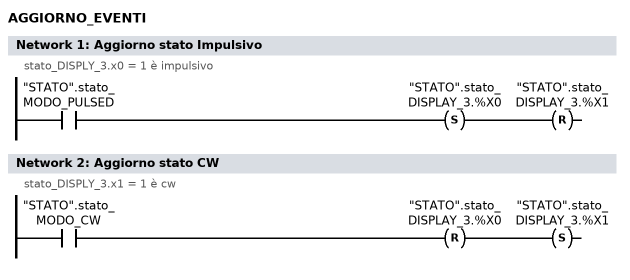
   RUNG wire#powerrail
      Contact( "STATO".stato_MODO_PULSED )
      S_Coil( "STATO".stato_DISPLAY_3.%X0 )
      R_Coil( "STATO".stato_DISPLAY_3.%X1 )
   END_RUNG
   // the same network as SCL:
   IF "STATO".stato_MODO_PULSED THEN
       "STATO".stato_DISPLAY_3.%X0 := TRUE;
       "STATO".stato_DISPLAY_3.%X1 := FALSE;
   END_IF;
END_REGION

REGION Network 2: Aggiorno stato CW
   // stato_DISPLY_3.x1 = 1 è cw
   RUNG wire#powerrail
      Contact( "STATO".stato_MODO_CW )
      R_Coil( "STATO".stato_DISPLAY_3.%X0 )
      S_Coil( "STATO".stato_DISPLAY_3.%X1 )
   END_RUNG
   // the same network as SCL:
   IF "STATO".stato_MODO_CW THEN
       "STATO".stato_DISPLAY_3.%X0 := FALSE;
       "STATO".stato_DISPLAY_3.%X1 := TRUE;
   END_IF;
END_REGION
END_FUNCTION

FUNCTION "LINEARIZZA_POTENZA" : Void   // FC11, LAD
TITLE = LINEARIZZA POTENZA
{ S7_Optimized_Access := 'FALSE' }
VERSION : 0.1
// Funzione di linearizzazione della potenza FWD e REFL
   VAR_TEMP   // added for the SCL form of the ladder/FBD networks
      _w1 : Bool;
   END_VAR
BEGIN

REGION Network 1: Calcolo indici N e N+1 tabella e punto adc&31
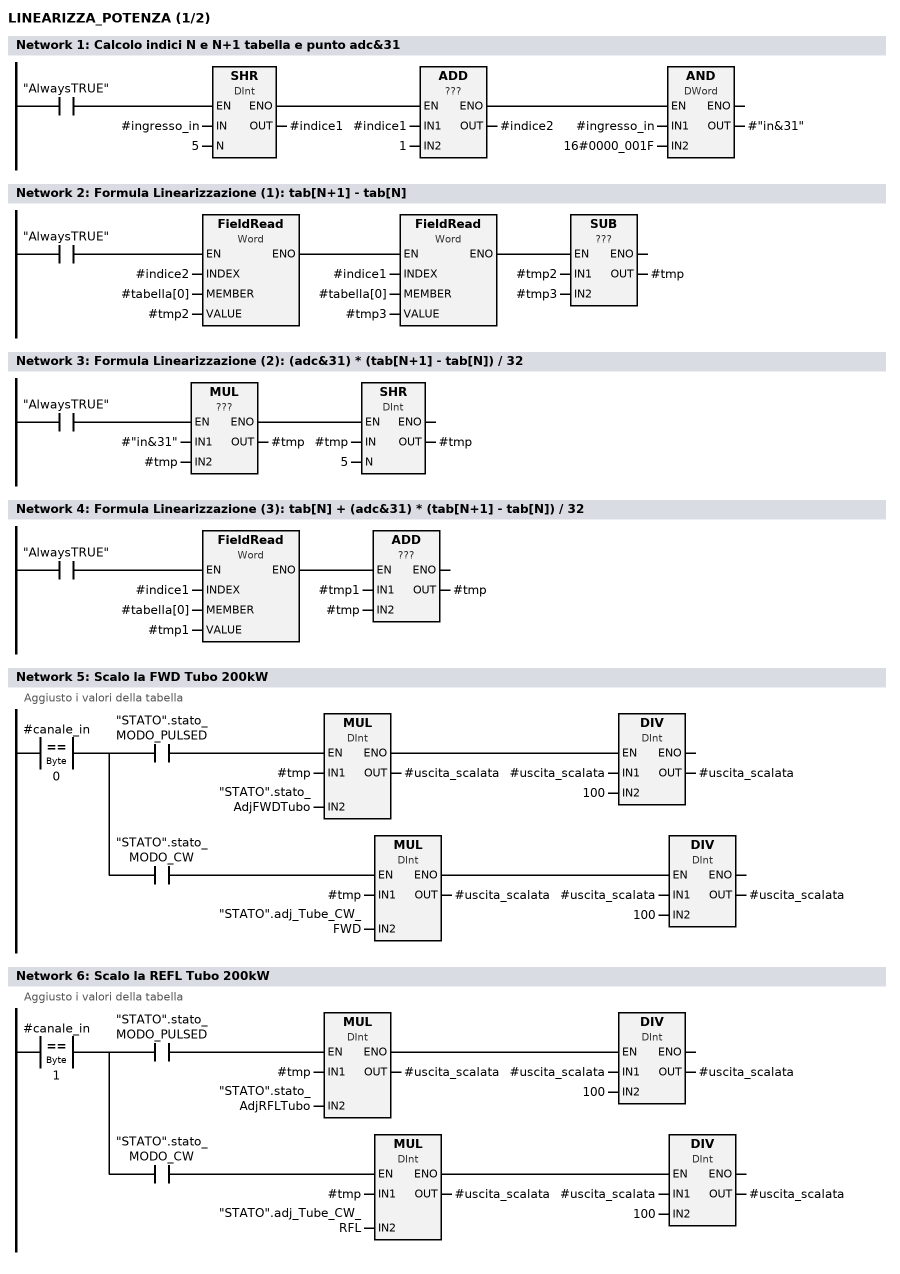
   // no checked SCL form for this network; see the picture
END_REGION

REGION Network 2: Formula Linearizzazione (1): tab[N+1] - tab[N]
   // no SCL statement known for FieldRead: written as a call
   // ENO of a box is taken as its EN; it also drops when the box reports an error
   #_w1 := "AlwaysTRUE";
   IF #_w1 THEN
       FieldRead(index := #indice2, member := #tabella[0], value := #tmp2);
       FieldRead(index := #indice1, member := #tabella[0], value := #tmp3);
       #tmp := #tmp2 - #tmp3;
   END_IF;
END_REGION

REGION Network 3: Formula Linearizzazione (2): (adc&31) * (tab[N+1] - tab[N]) / 32
   RUNG wire#powerrail
      Contact( "AlwaysTRUE" )
      { S7_Templates := "SrcType := ???" } Mul(in1 := #"in&31", in2 := #tmp, out => #tmp)
      { S7_Templates := "SrcType := DInt" } Shr(in := #tmp, n := 5, out => #tmp)
   END_RUNG
   // the same network as SCL:
   IF "AlwaysTRUE" THEN
       #tmp := #"in&31" * #tmp;
       #tmp := SHR(IN := #tmp, N := 5);
   END_IF;
END_REGION

REGION Network 4: Formula Linearizzazione (3): tab[N] + (adc&31) * (tab[N+1] - tab[N]) / 32
   // no SCL statement known for FieldRead: written as a call
   // ENO of a box is taken as its EN; it also drops when the box reports an error
   #_w1 := "AlwaysTRUE";
   IF #_w1 THEN
       FieldRead(index := #indice1, member := #tabella[0], value := #tmp1);
       #tmp := #tmp1 + #tmp;
   END_IF;
END_REGION

REGION Network 5: Scalo la FWD Tubo 200kW
   // Aggiusto i valori della tabella
   RUNG wire#powerrail
      { S7_Templates := "SrcType := Byte" } EQ_Contact(in1 := #canale_in, in2 := 0)
      wire#w1
      Contact( "STATO".stato_MODO_PULSED )
      { S7_Templates := "SrcType := DInt" } Mul(in1 := #tmp, in2 := "STATO".stato_AdjFWDTubo, out => #uscita_scalata)
      { S7_Templates := "SrcType := DInt" } Div(in1 := #uscita_scalata, in2 := 100, out => #uscita_scalata)
   END_RUNG
   RUNG wire#w1
      Contact( "STATO".stato_MODO_CW )
      { S7_Templates := "SrcType := DInt" } Mul(in1 := #tmp, in2 := "STATO".adj_Tube_CW_FWD, out => #uscita_scalata)
      { S7_Templates := "SrcType := DInt" } Div(in1 := #uscita_scalata, in2 := 100, out => #uscita_scalata)
   END_RUNG
   // the same network as SCL:
   #_w1 := #canale_in = 0;
   IF #_w1 AND "STATO".stato_MODO_PULSED THEN
       #uscita_scalata := #tmp * "STATO".stato_AdjFWDTubo;
       #uscita_scalata := #uscita_scalata / 100;
   END_IF;
   IF #_w1 AND "STATO".stato_MODO_CW THEN
       #uscita_scalata := #tmp * "STATO".adj_Tube_CW_FWD;
       #uscita_scalata := #uscita_scalata / 100;
   END_IF;
END_REGION

REGION Network 6: Scalo la REFL Tubo 200kW
   // Aggiusto i valori della tabella
   RUNG wire#powerrail
      { S7_Templates := "SrcType := Byte" } EQ_Contact(in1 := #canale_in, in2 := 1)
      wire#w1
      Contact( "STATO".stato_MODO_PULSED )
      { S7_Templates := "SrcType := DInt" } Mul(in1 := #tmp, in2 := "STATO".stato_AdjRFLTubo, out => #uscita_scalata)
      { S7_Templates := "SrcType := DInt" } Div(in1 := #uscita_scalata, in2 := 100, out => #uscita_scalata)
   END_RUNG
   RUNG wire#w1
      Contact( "STATO".stato_MODO_CW )
      { S7_Templates := "SrcType := DInt" } Mul(in1 := #tmp, in2 := "STATO".adj_Tube_CW_RFL, out => #uscita_scalata)
      { S7_Templates := "SrcType := DInt" } Div(in1 := #uscita_scalata, in2 := 100, out => #uscita_scalata)
   END_RUNG
   // the same network as SCL:
   #_w1 := #canale_in = 1;
   IF #_w1 AND "STATO".stato_MODO_PULSED THEN
       #uscita_scalata := #tmp * "STATO".stato_AdjRFLTubo;
       #uscita_scalata := #uscita_scalata / 100;
   END_IF;
   IF #_w1 AND "STATO".stato_MODO_CW THEN
       #uscita_scalata := #tmp * "STATO".adj_Tube_CW_RFL;
       #uscita_scalata := #uscita_scalata / 100;
   END_IF;
END_REGION

REGION Network 7: Scalo la FWD Stato Solido
   // Aggiusto i valori della tabella
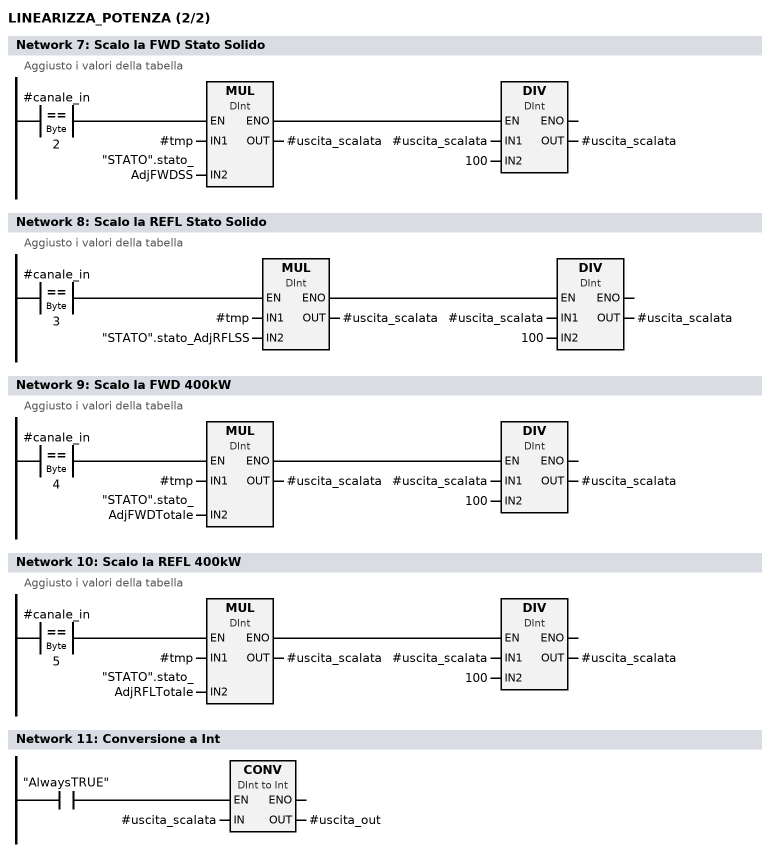
   RUNG wire#powerrail
      { S7_Templates := "SrcType := Byte" } EQ_Contact(in1 := #canale_in, in2 := 2)
      { S7_Templates := "SrcType := DInt" } Mul(in1 := #tmp, in2 := "STATO".stato_AdjFWDSS, out => #uscita_scalata)
      { S7_Templates := "SrcType := DInt" } Div(in1 := #uscita_scalata, in2 := 100, out => #uscita_scalata)
   END_RUNG
   // the same network as SCL:
   IF #canale_in = 2 THEN
       #uscita_scalata := #tmp * "STATO".stato_AdjFWDSS;
       #uscita_scalata := #uscita_scalata / 100;
   END_IF;
END_REGION

REGION Network 8: Scalo la REFL Stato Solido
   // Aggiusto i valori della tabella
   RUNG wire#powerrail
      { S7_Templates := "SrcType := Byte" } EQ_Contact(in1 := #canale_in, in2 := 3)
      { S7_Templates := "SrcType := DInt" } Mul(in1 := #tmp, in2 := "STATO".stato_AdjRFLSS, out => #uscita_scalata)
      { S7_Templates := "SrcType := DInt" } Div(in1 := #uscita_scalata, in2 := 100, out => #uscita_scalata)
   END_RUNG
   // the same network as SCL:
   IF #canale_in = 3 THEN
       #uscita_scalata := #tmp * "STATO".stato_AdjRFLSS;
       #uscita_scalata := #uscita_scalata / 100;
   END_IF;
END_REGION

REGION Network 9: Scalo la FWD 400kW
   // Aggiusto i valori della tabella
   RUNG wire#powerrail
      { S7_Templates := "SrcType := Byte" } EQ_Contact(in1 := #canale_in, in2 := 4)
      { S7_Templates := "SrcType := DInt" } Mul(in1 := #tmp, in2 := "STATO".stato_AdjFWDTotale, out => #uscita_scalata)
      { S7_Templates := "SrcType := DInt" } Div(in1 := #uscita_scalata, in2 := 100, out => #uscita_scalata)
   END_RUNG
   // the same network as SCL:
   IF #canale_in = 4 THEN
       #uscita_scalata := #tmp * "STATO".stato_AdjFWDTotale;
       #uscita_scalata := #uscita_scalata / 100;
   END_IF;
END_REGION

REGION Network 10: Scalo la REFL 400kW
   // Aggiusto i valori della tabella
   RUNG wire#powerrail
      { S7_Templates := "SrcType := Byte" } EQ_Contact(in1 := #canale_in, in2 := 5)
      { S7_Templates := "SrcType := DInt" } Mul(in1 := #tmp, in2 := "STATO".stato_AdjRFLTotale, out => #uscita_scalata)
      { S7_Templates := "SrcType := DInt" } Div(in1 := #uscita_scalata, in2 := 100, out => #uscita_scalata)
   END_RUNG
   // the same network as SCL:
   IF #canale_in = 5 THEN
       #uscita_scalata := #tmp * "STATO".stato_AdjRFLTotale;
       #uscita_scalata := #uscita_scalata / 100;
   END_IF;
END_REGION

REGION Network 11: Conversione a Int
   RUNG wire#powerrail
      Contact( "AlwaysTRUE" )
      { S7_Templates := "[SrcType := DInt, DestType := Int]" } Convert(in := #uscita_scalata, out => #uscita_out)
   END_RUNG
   // the same network as SCL:
   IF "AlwaysTRUE" THEN #uscita_out := DINT_TO_INT(#uscita_scalata); END_IF;
END_REGION
END_FUNCTION

FUNCTION "TRADUCI_TLS" : Void   // FC12, LAD
TITLE = TRADUCI_TLS
{ S7_Optimized_Access := 'FALSE' }
VERSION : 0.1
// Traduce gli stati/allarmi/misure in formato DATABLOCCO (EPICS_READ DB27) per l'invio al partner remoto EPICS.
   VAR_TEMP   // added for the SCL form of the ladder/FBD networks
      _w1 : Bool;
   END_VAR
BEGIN

REGION Network 1: Stato Locale/Remoto
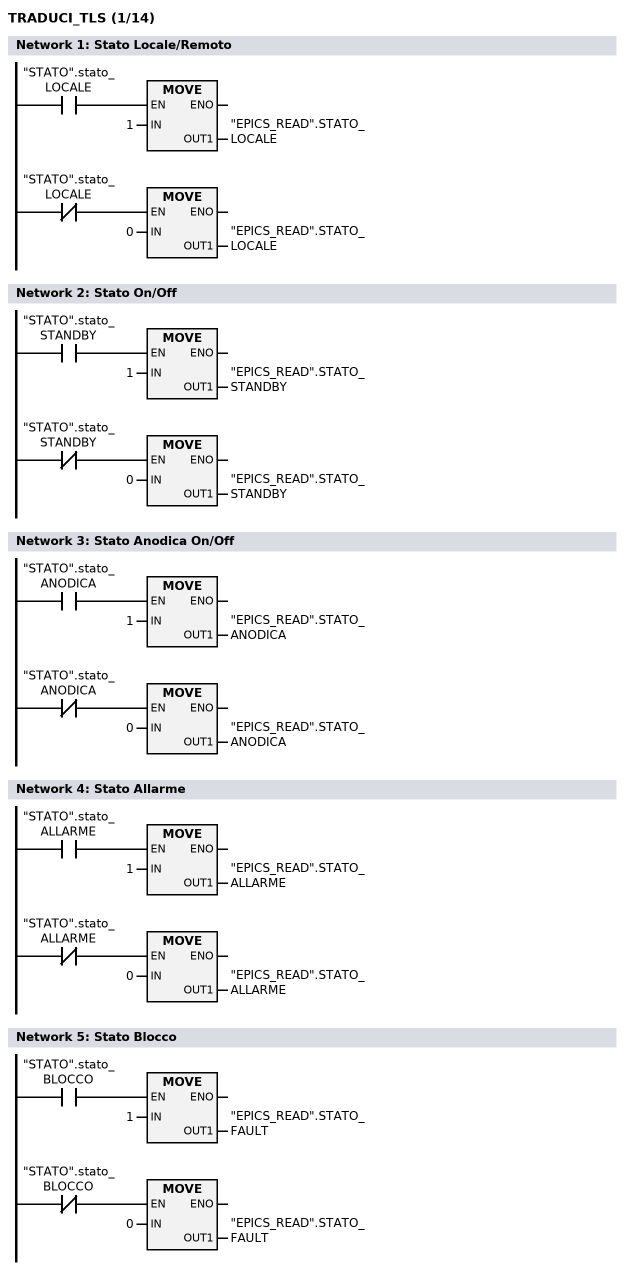
   RUNG wire#powerrail
      Contact( "STATO".stato_LOCALE )
      Move(in := 1, out1 => "EPICS_READ".STATO_LOCALE)
   END_RUNG
   RUNG wire#powerrail
      I_Contact( "STATO".stato_LOCALE )
      Move(in := 0, out1 => "EPICS_READ".STATO_LOCALE)
   END_RUNG
   // the same network as SCL:
   IF "STATO".stato_LOCALE THEN "EPICS_READ".STATO_LOCALE := 1; END_IF;
   IF NOT "STATO".stato_LOCALE THEN "EPICS_READ".STATO_LOCALE := 0; END_IF;
END_REGION

REGION Network 2: Stato On/Off
   RUNG wire#powerrail
      Contact( "STATO".stato_STANDBY )
      Move(in := 1, out1 => "EPICS_READ".STATO_STANDBY)
   END_RUNG
   RUNG wire#powerrail
      I_Contact( "STATO".stato_STANDBY )
      Move(in := 0, out1 => "EPICS_READ".STATO_STANDBY)
   END_RUNG
   // the same network as SCL:
   IF "STATO".stato_STANDBY THEN "EPICS_READ".STATO_STANDBY := 1; END_IF;
   IF NOT "STATO".stato_STANDBY THEN "EPICS_READ".STATO_STANDBY := 0; END_IF;
END_REGION

REGION Network 3: Stato Anodica On/Off
   RUNG wire#powerrail
      Contact( "STATO".stato_ANODICA )
      Move(in := 1, out1 => "EPICS_READ".STATO_ANODICA)
   END_RUNG
   RUNG wire#powerrail
      I_Contact( "STATO".stato_ANODICA )
      Move(in := 0, out1 => "EPICS_READ".STATO_ANODICA)
   END_RUNG
   // the same network as SCL:
   IF "STATO".stato_ANODICA THEN "EPICS_READ".STATO_ANODICA := 1; END_IF;
   IF NOT "STATO".stato_ANODICA THEN "EPICS_READ".STATO_ANODICA := 0; END_IF;
END_REGION

REGION Network 4: Stato Allarme
   RUNG wire#powerrail
      Contact( "STATO".stato_ALLARME )
      Move(in := 1, out1 => "EPICS_READ".STATO_ALLARME)
   END_RUNG
   RUNG wire#powerrail
      I_Contact( "STATO".stato_ALLARME )
      Move(in := 0, out1 => "EPICS_READ".STATO_ALLARME)
   END_RUNG
   // the same network as SCL:
   IF "STATO".stato_ALLARME THEN "EPICS_READ".STATO_ALLARME := 1; END_IF;
   IF NOT "STATO".stato_ALLARME THEN "EPICS_READ".STATO_ALLARME := 0; END_IF;
END_REGION

REGION Network 5: Stato Blocco
   RUNG wire#powerrail
      Contact( "STATO".stato_BLOCCO )
      Move(in := 1, out1 => "EPICS_READ".STATO_FAULT)
   END_RUNG
   RUNG wire#powerrail
      I_Contact( "STATO".stato_BLOCCO )
      Move(in := 0, out1 => "EPICS_READ".STATO_FAULT)
   END_RUNG
   // the same network as SCL:
   IF "STATO".stato_BLOCCO THEN "EPICS_READ".STATO_FAULT := 1; END_IF;
   IF NOT "STATO".stato_BLOCCO THEN "EPICS_READ".STATO_FAULT := 0; END_IF;
END_REGION

REGION Network 6: Impulsivo/CW
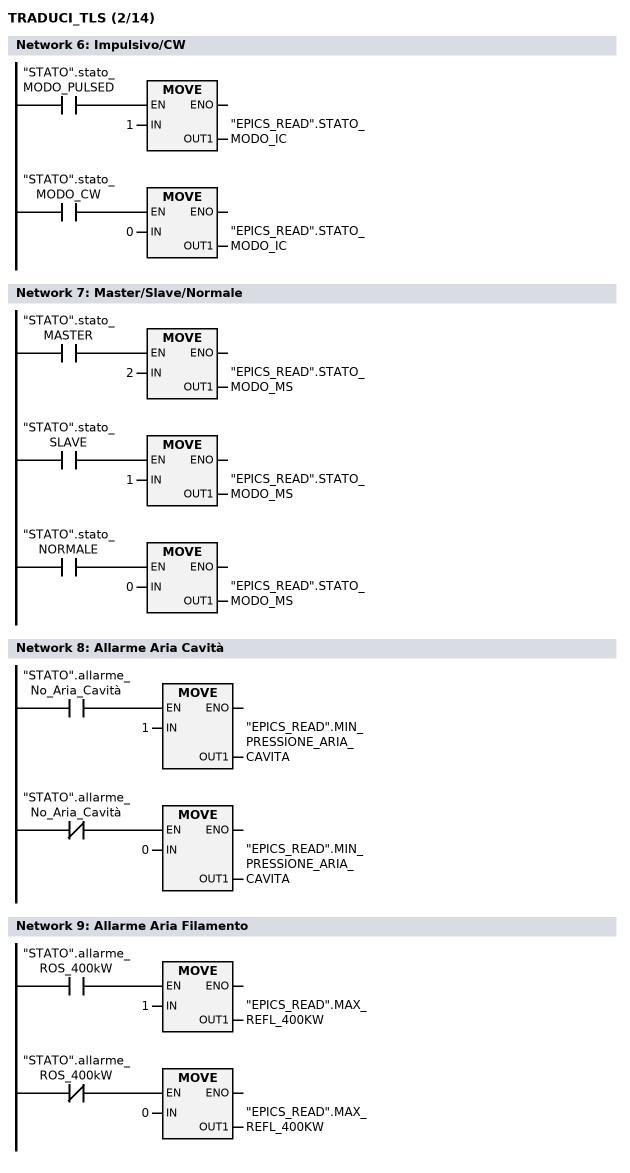
   RUNG wire#powerrail
      Contact( "STATO".stato_MODO_PULSED )
      Move(in := 1, out1 => "EPICS_READ".STATO_MODO_IC)
   END_RUNG
   RUNG wire#powerrail
      Contact( "STATO".stato_MODO_CW )
      Move(in := 0, out1 => "EPICS_READ".STATO_MODO_IC)
   END_RUNG
   // the same network as SCL:
   IF "STATO".stato_MODO_PULSED THEN "EPICS_READ".STATO_MODO_IC := 1; END_IF;
   IF "STATO".stato_MODO_CW THEN "EPICS_READ".STATO_MODO_IC := 0; END_IF;
END_REGION

REGION Network 7: Master/Slave/Normale
   RUNG wire#powerrail
      Contact( "STATO".stato_MASTER )
      Move(in := 2, out1 => "EPICS_READ".STATO_MODO_MS)
   END_RUNG
   RUNG wire#powerrail
      Contact( "STATO".stato_SLAVE )
      Move(in := 1, out1 => "EPICS_READ".STATO_MODO_MS)
   END_RUNG
   RUNG wire#powerrail
      Contact( "STATO".stato_NORMALE )
      Move(in := 0, out1 => "EPICS_READ".STATO_MODO_MS)
   END_RUNG
   // the same network as SCL:
   IF "STATO".stato_MASTER THEN "EPICS_READ".STATO_MODO_MS := 2; END_IF;
   IF "STATO".stato_SLAVE THEN "EPICS_READ".STATO_MODO_MS := 1; END_IF;
   IF "STATO".stato_NORMALE THEN "EPICS_READ".STATO_MODO_MS := 0; END_IF;
END_REGION

REGION Network 8: Allarme Aria Cavità
   RUNG wire#powerrail
      Contact( "STATO".allarme_No_Aria_Cavità )
      Move(in := 1, out1 => "EPICS_READ".MIN_PRESSIONE_ARIA_CAVITA)
   END_RUNG
   RUNG wire#powerrail
      I_Contact( "STATO".allarme_No_Aria_Cavità )
      Move(in := 0, out1 => "EPICS_READ".MIN_PRESSIONE_ARIA_CAVITA)
   END_RUNG
   // the same network as SCL:
   IF "STATO".allarme_No_Aria_Cavità THEN "EPICS_READ".MIN_PRESSIONE_ARIA_CAVITA := 1; END_IF;
   IF NOT "STATO".allarme_No_Aria_Cavità THEN "EPICS_READ".MIN_PRESSIONE_ARIA_CAVITA := 0; END_IF;
END_REGION

REGION Network 9: Allarme Aria Filamento
   RUNG wire#powerrail
      Contact( "STATO".allarme_ROS_400kW )
      Move(in := 1, out1 => "EPICS_READ".MAX_REFL_400KW)
   END_RUNG
   RUNG wire#powerrail
      I_Contact( "STATO".allarme_ROS_400kW )
      Move(in := 0, out1 => "EPICS_READ".MAX_REFL_400KW)
   END_RUNG
   // the same network as SCL:
   IF "STATO".allarme_ROS_400kW THEN "EPICS_READ".MAX_REFL_400KW := 1; END_IF;
   IF NOT "STATO".allarme_ROS_400kW THEN "EPICS_READ".MAX_REFL_400KW := 0; END_IF;
END_REGION

REGION Network 10: Allarme Flusso LQD Tubo
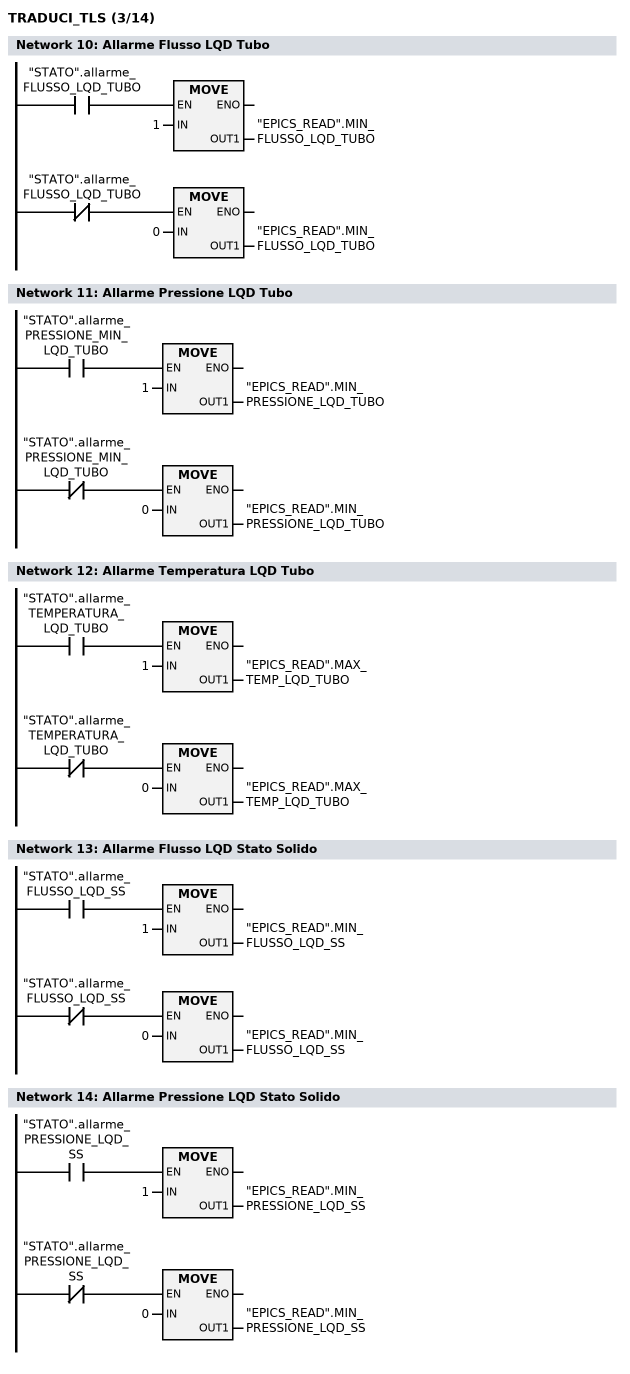
   RUNG wire#powerrail
      Contact( "STATO".allarme_FLUSSO_LQD_TUBO )
      Move(in := 1, out1 => "EPICS_READ".MIN_FLUSSO_LQD_TUBO)
   END_RUNG
   RUNG wire#powerrail
      I_Contact( "STATO".allarme_FLUSSO_LQD_TUBO )
      Move(in := 0, out1 => "EPICS_READ".MIN_FLUSSO_LQD_TUBO)
   END_RUNG
   // the same network as SCL:
   IF "STATO".allarme_FLUSSO_LQD_TUBO THEN "EPICS_READ".MIN_FLUSSO_LQD_TUBO := 1; END_IF;
   IF NOT "STATO".allarme_FLUSSO_LQD_TUBO THEN "EPICS_READ".MIN_FLUSSO_LQD_TUBO := 0; END_IF;
END_REGION

REGION Network 11: Allarme Pressione LQD Tubo
   RUNG wire#powerrail
      Contact( "STATO".allarme_PRESSIONE_MIN_LQD_TUBO )
      Move(in := 1, out1 => "EPICS_READ".MIN_PRESSIONE_LQD_TUBO)
   END_RUNG
   RUNG wire#powerrail
      I_Contact( "STATO".allarme_PRESSIONE_MIN_LQD_TUBO )
      Move(in := 0, out1 => "EPICS_READ".MIN_PRESSIONE_LQD_TUBO)
   END_RUNG
   // the same network as SCL:
   IF "STATO".allarme_PRESSIONE_MIN_LQD_TUBO THEN "EPICS_READ".MIN_PRESSIONE_LQD_TUBO := 1; END_IF;
   IF NOT "STATO".allarme_PRESSIONE_MIN_LQD_TUBO THEN "EPICS_READ".MIN_PRESSIONE_LQD_TUBO := 0; END_IF;
END_REGION

REGION Network 12: Allarme Temperatura LQD Tubo
   RUNG wire#powerrail
      Contact( "STATO".allarme_TEMPERATURA_LQD_TUBO )
      Move(in := 1, out1 => "EPICS_READ".MAX_TEMP_LQD_TUBO)
   END_RUNG
   RUNG wire#powerrail
      I_Contact( "STATO".allarme_TEMPERATURA_LQD_TUBO )
      Move(in := 0, out1 => "EPICS_READ".MAX_TEMP_LQD_TUBO)
   END_RUNG
   // the same network as SCL:
   IF "STATO".allarme_TEMPERATURA_LQD_TUBO THEN "EPICS_READ".MAX_TEMP_LQD_TUBO := 1; END_IF;
   IF NOT "STATO".allarme_TEMPERATURA_LQD_TUBO THEN "EPICS_READ".MAX_TEMP_LQD_TUBO := 0; END_IF;
END_REGION

REGION Network 13: Allarme Flusso LQD Stato Solido
   RUNG wire#powerrail
      Contact( "STATO".allarme_FLUSSO_LQD_SS )
      Move(in := 1, out1 => "EPICS_READ".MIN_FLUSSO_LQD_SS)
   END_RUNG
   RUNG wire#powerrail
      I_Contact( "STATO".allarme_FLUSSO_LQD_SS )
      Move(in := 0, out1 => "EPICS_READ".MIN_FLUSSO_LQD_SS)
   END_RUNG
   // the same network as SCL:
   IF "STATO".allarme_FLUSSO_LQD_SS THEN "EPICS_READ".MIN_FLUSSO_LQD_SS := 1; END_IF;
   IF NOT "STATO".allarme_FLUSSO_LQD_SS THEN "EPICS_READ".MIN_FLUSSO_LQD_SS := 0; END_IF;
END_REGION

REGION Network 14: Allarme Pressione LQD Stato Solido
   RUNG wire#powerrail
      Contact( "STATO".allarme_PRESSIONE_LQD_SS )
      Move(in := 1, out1 => "EPICS_READ".MIN_PRESSIONE_LQD_SS)
   END_RUNG
   RUNG wire#powerrail
      I_Contact( "STATO".allarme_PRESSIONE_LQD_SS )
      Move(in := 0, out1 => "EPICS_READ".MIN_PRESSIONE_LQD_SS)
   END_RUNG
   // the same network as SCL:
   IF "STATO".allarme_PRESSIONE_LQD_SS THEN "EPICS_READ".MIN_PRESSIONE_LQD_SS := 1; END_IF;
   IF NOT "STATO".allarme_PRESSIONE_LQD_SS THEN "EPICS_READ".MIN_PRESSIONE_LQD_SS := 0; END_IF;
END_REGION

REGION Network 15: Allarme Temperatura LQD Stato Solido
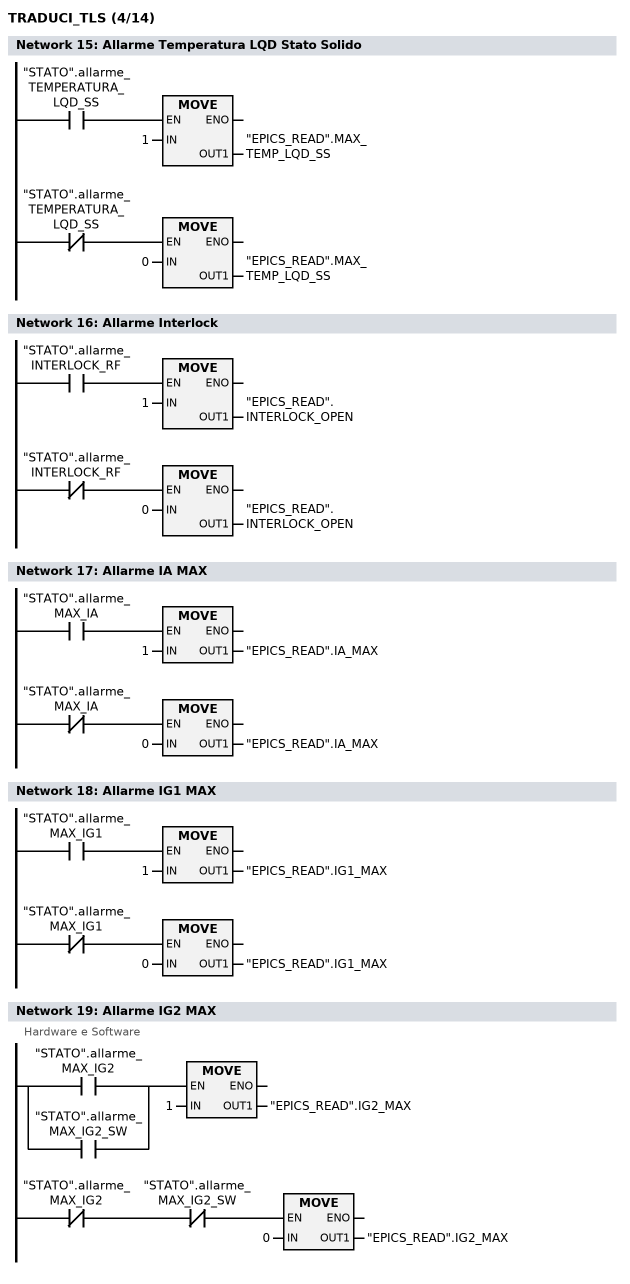
   RUNG wire#powerrail
      Contact( "STATO".allarme_TEMPERATURA_LQD_SS )
      Move(in := 1, out1 => "EPICS_READ".MAX_TEMP_LQD_SS)
   END_RUNG
   RUNG wire#powerrail
      I_Contact( "STATO".allarme_TEMPERATURA_LQD_SS )
      Move(in := 0, out1 => "EPICS_READ".MAX_TEMP_LQD_SS)
   END_RUNG
   // the same network as SCL:
   IF "STATO".allarme_TEMPERATURA_LQD_SS THEN "EPICS_READ".MAX_TEMP_LQD_SS := 1; END_IF;
   IF NOT "STATO".allarme_TEMPERATURA_LQD_SS THEN "EPICS_READ".MAX_TEMP_LQD_SS := 0; END_IF;
END_REGION

REGION Network 16: Allarme Interlock
   RUNG wire#powerrail
      Contact( "STATO".allarme_INTERLOCK_RF )
      Move(in := 1, out1 => "EPICS_READ".INTERLOCK_OPEN)
   END_RUNG
   RUNG wire#powerrail
      I_Contact( "STATO".allarme_INTERLOCK_RF )
      Move(in := 0, out1 => "EPICS_READ".INTERLOCK_OPEN)
   END_RUNG
   // the same network as SCL:
   IF "STATO".allarme_INTERLOCK_RF THEN "EPICS_READ".INTERLOCK_OPEN := 1; END_IF;
   IF NOT "STATO".allarme_INTERLOCK_RF THEN "EPICS_READ".INTERLOCK_OPEN := 0; END_IF;
END_REGION

REGION Network 17: Allarme IA MAX
   RUNG wire#powerrail
      Contact( "STATO".allarme_MAX_IA )
      Move(in := 1, out1 => "EPICS_READ".IA_MAX)
   END_RUNG
   RUNG wire#powerrail
      I_Contact( "STATO".allarme_MAX_IA )
      Move(in := 0, out1 => "EPICS_READ".IA_MAX)
   END_RUNG
   // the same network as SCL:
   IF "STATO".allarme_MAX_IA THEN "EPICS_READ".IA_MAX := 1; END_IF;
   IF NOT "STATO".allarme_MAX_IA THEN "EPICS_READ".IA_MAX := 0; END_IF;
END_REGION

REGION Network 18: Allarme IG1 MAX
   RUNG wire#powerrail
      Contact( "STATO".allarme_MAX_IG1 )
      Move(in := 1, out1 => "EPICS_READ".IG1_MAX)
   END_RUNG
   RUNG wire#powerrail
      I_Contact( "STATO".allarme_MAX_IG1 )
      Move(in := 0, out1 => "EPICS_READ".IG1_MAX)
   END_RUNG
   // the same network as SCL:
   IF "STATO".allarme_MAX_IG1 THEN "EPICS_READ".IG1_MAX := 1; END_IF;
   IF NOT "STATO".allarme_MAX_IG1 THEN "EPICS_READ".IG1_MAX := 0; END_IF;
END_REGION

REGION Network 19: Allarme IG2 MAX
   // Hardware e Software
   RUNG wire#powerrail
      Contact( "STATO".allarme_MAX_IG2 )
      wire#w1
      Move(in := 1, out1 => "EPICS_READ".IG2_MAX)
   END_RUNG
   RUNG wire#powerrail
      Contact( "STATO".allarme_MAX_IG2_SW )
   END_RUNG wire#w1
   RUNG wire#powerrail
      I_Contact( "STATO".allarme_MAX_IG2 )
      I_Contact( "STATO".allarme_MAX_IG2_SW )
      Move(in := 0, out1 => "EPICS_READ".IG2_MAX)
   END_RUNG
   // the same network as SCL:
   IF "STATO".allarme_MAX_IG2 OR "STATO".allarme_MAX_IG2_SW THEN "EPICS_READ".IG2_MAX := 1; END_IF;
   IF NOT "STATO".allarme_MAX_IG2 AND NOT "STATO".allarme_MAX_IG2_SW THEN "EPICS_READ".IG2_MAX := 0; END_IF;
END_REGION

REGION Network 20: Allarme Crowbar
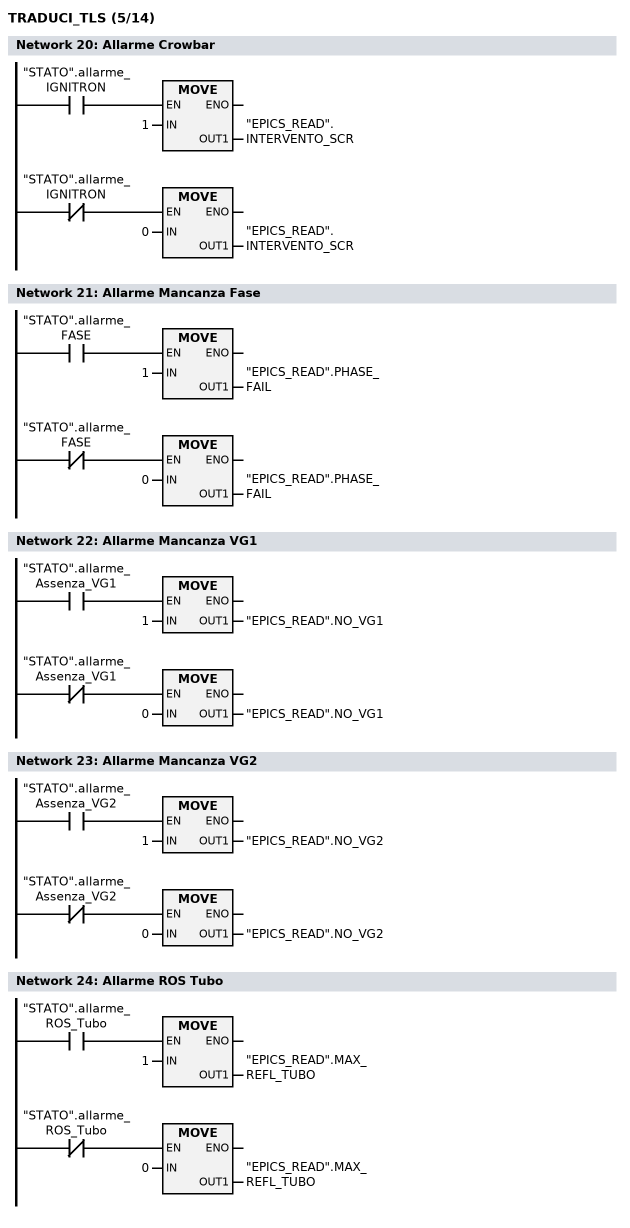
   RUNG wire#powerrail
      Contact( "STATO".allarme_IGNITRON )
      Move(in := 1, out1 => "EPICS_READ".INTERVENTO_SCR)
   END_RUNG
   RUNG wire#powerrail
      I_Contact( "STATO".allarme_IGNITRON )
      Move(in := 0, out1 => "EPICS_READ".INTERVENTO_SCR)
   END_RUNG
   // the same network as SCL:
   IF "STATO".allarme_IGNITRON THEN "EPICS_READ".INTERVENTO_SCR := 1; END_IF;
   IF NOT "STATO".allarme_IGNITRON THEN "EPICS_READ".INTERVENTO_SCR := 0; END_IF;
END_REGION

REGION Network 21: Allarme Mancanza Fase
   RUNG wire#powerrail
      Contact( "STATO".allarme_FASE )
      Move(in := 1, out1 => "EPICS_READ".PHASE_FAIL)
   END_RUNG
   RUNG wire#powerrail
      I_Contact( "STATO".allarme_FASE )
      Move(in := 0, out1 => "EPICS_READ".PHASE_FAIL)
   END_RUNG
   // the same network as SCL:
   IF "STATO".allarme_FASE THEN "EPICS_READ".PHASE_FAIL := 1; END_IF;
   IF NOT "STATO".allarme_FASE THEN "EPICS_READ".PHASE_FAIL := 0; END_IF;
END_REGION

REGION Network 22: Allarme Mancanza VG1
   RUNG wire#powerrail
      Contact( "STATO".allarme_Assenza_VG1 )
      Move(in := 1, out1 => "EPICS_READ".NO_VG1)
   END_RUNG
   RUNG wire#powerrail
      I_Contact( "STATO".allarme_Assenza_VG1 )
      Move(in := 0, out1 => "EPICS_READ".NO_VG1)
   END_RUNG
   // the same network as SCL:
   IF "STATO".allarme_Assenza_VG1 THEN "EPICS_READ".NO_VG1 := 1; END_IF;
   IF NOT "STATO".allarme_Assenza_VG1 THEN "EPICS_READ".NO_VG1 := 0; END_IF;
END_REGION

REGION Network 23: Allarme Mancanza VG2
   RUNG wire#powerrail
      Contact( "STATO".allarme_Assenza_VG2 )
      Move(in := 1, out1 => "EPICS_READ".NO_VG2)
   END_RUNG
   RUNG wire#powerrail
      I_Contact( "STATO".allarme_Assenza_VG2 )
      Move(in := 0, out1 => "EPICS_READ".NO_VG2)
   END_RUNG
   // the same network as SCL:
   IF "STATO".allarme_Assenza_VG2 THEN "EPICS_READ".NO_VG2 := 1; END_IF;
   IF NOT "STATO".allarme_Assenza_VG2 THEN "EPICS_READ".NO_VG2 := 0; END_IF;
END_REGION

REGION Network 24: Allarme ROS Tubo
   RUNG wire#powerrail
      Contact( "STATO".allarme_ROS_Tubo )
      Move(in := 1, out1 => "EPICS_READ".MAX_REFL_TUBO)
   END_RUNG
   RUNG wire#powerrail
      I_Contact( "STATO".allarme_ROS_Tubo )
      Move(in := 0, out1 => "EPICS_READ".MAX_REFL_TUBO)
   END_RUNG
   // the same network as SCL:
   IF "STATO".allarme_ROS_Tubo THEN "EPICS_READ".MAX_REFL_TUBO := 1; END_IF;
   IF NOT "STATO".allarme_ROS_Tubo THEN "EPICS_READ".MAX_REFL_TUBO := 0; END_IF;
END_REGION

REGION Network 25: Allarme ROS Stato Solido
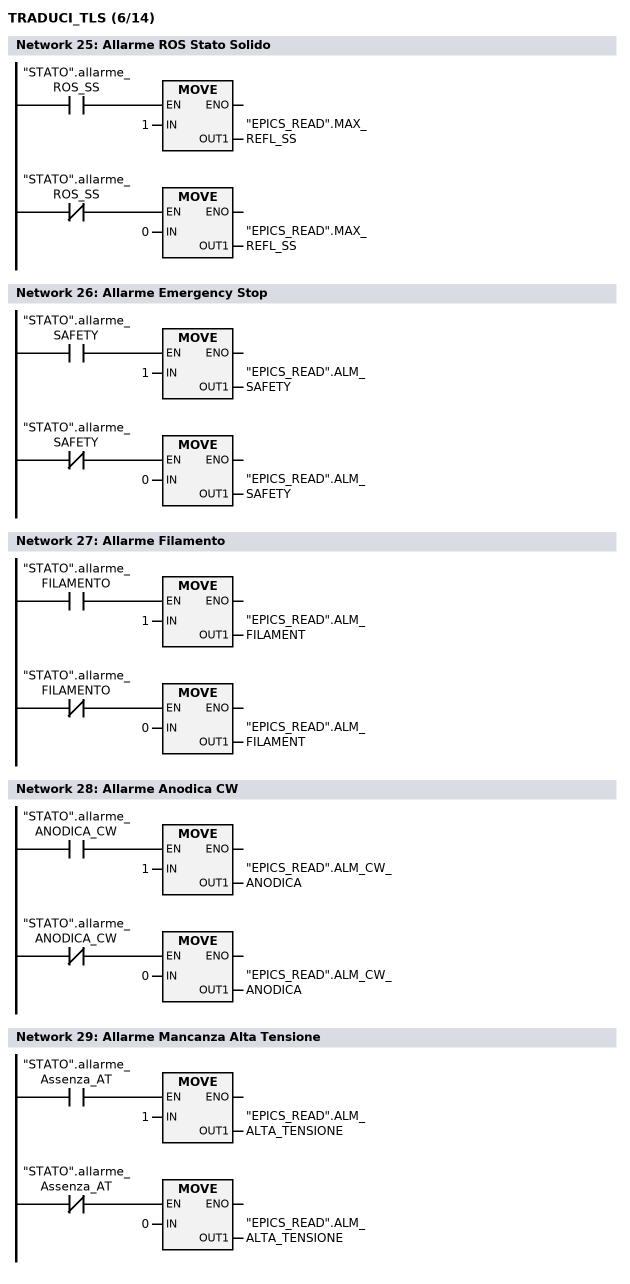
   RUNG wire#powerrail
      Contact( "STATO".allarme_ROS_SS )
      Move(in := 1, out1 => "EPICS_READ".MAX_REFL_SS)
   END_RUNG
   RUNG wire#powerrail
      I_Contact( "STATO".allarme_ROS_SS )
      Move(in := 0, out1 => "EPICS_READ".MAX_REFL_SS)
   END_RUNG
   // the same network as SCL:
   IF "STATO".allarme_ROS_SS THEN "EPICS_READ".MAX_REFL_SS := 1; END_IF;
   IF NOT "STATO".allarme_ROS_SS THEN "EPICS_READ".MAX_REFL_SS := 0; END_IF;
END_REGION

REGION Network 26: Allarme Emergency Stop
   RUNG wire#powerrail
      Contact( "STATO".allarme_SAFETY )
      Move(in := 1, out1 => "EPICS_READ".ALM_SAFETY)
   END_RUNG
   RUNG wire#powerrail
      I_Contact( "STATO".allarme_SAFETY )
      Move(in := 0, out1 => "EPICS_READ".ALM_SAFETY)
   END_RUNG
   // the same network as SCL:
   IF "STATO".allarme_SAFETY THEN "EPICS_READ".ALM_SAFETY := 1; END_IF;
   IF NOT "STATO".allarme_SAFETY THEN "EPICS_READ".ALM_SAFETY := 0; END_IF;
END_REGION

REGION Network 27: Allarme Filamento
   RUNG wire#powerrail
      Contact( "STATO".allarme_FILAMENTO )
      Move(in := 1, out1 => "EPICS_READ".ALM_FILAMENT)
   END_RUNG
   RUNG wire#powerrail
      I_Contact( "STATO".allarme_FILAMENTO )
      Move(in := 0, out1 => "EPICS_READ".ALM_FILAMENT)
   END_RUNG
   // the same network as SCL:
   IF "STATO".allarme_FILAMENTO THEN "EPICS_READ".ALM_FILAMENT := 1; END_IF;
   IF NOT "STATO".allarme_FILAMENTO THEN "EPICS_READ".ALM_FILAMENT := 0; END_IF;
END_REGION

REGION Network 28: Allarme Anodica CW
   RUNG wire#powerrail
      Contact( "STATO".allarme_ANODICA_CW )
      Move(in := 1, out1 => "EPICS_READ".ALM_CW_ANODICA)
   END_RUNG
   RUNG wire#powerrail
      I_Contact( "STATO".allarme_ANODICA_CW )
      Move(in := 0, out1 => "EPICS_READ".ALM_CW_ANODICA)
   END_RUNG
   // the same network as SCL:
   IF "STATO".allarme_ANODICA_CW THEN "EPICS_READ".ALM_CW_ANODICA := 1; END_IF;
   IF NOT "STATO".allarme_ANODICA_CW THEN "EPICS_READ".ALM_CW_ANODICA := 0; END_IF;
END_REGION

REGION Network 29: Allarme Mancanza Alta Tensione
   RUNG wire#powerrail
      Contact( "STATO".allarme_Assenza_AT )
      Move(in := 1, out1 => "EPICS_READ".ALM_ALTA_TENSIONE)
   END_RUNG
   RUNG wire#powerrail
      I_Contact( "STATO".allarme_Assenza_AT )
      Move(in := 0, out1 => "EPICS_READ".ALM_ALTA_TENSIONE)
   END_RUNG
   // the same network as SCL:
   IF "STATO".allarme_Assenza_AT THEN "EPICS_READ".ALM_ALTA_TENSIONE := 1; END_IF;
   IF NOT "STATO".allarme_Assenza_AT THEN "EPICS_READ".ALM_ALTA_TENSIONE := 0; END_IF;
END_REGION

REGION Network 30: Allarme Temperatura Alta Tensione
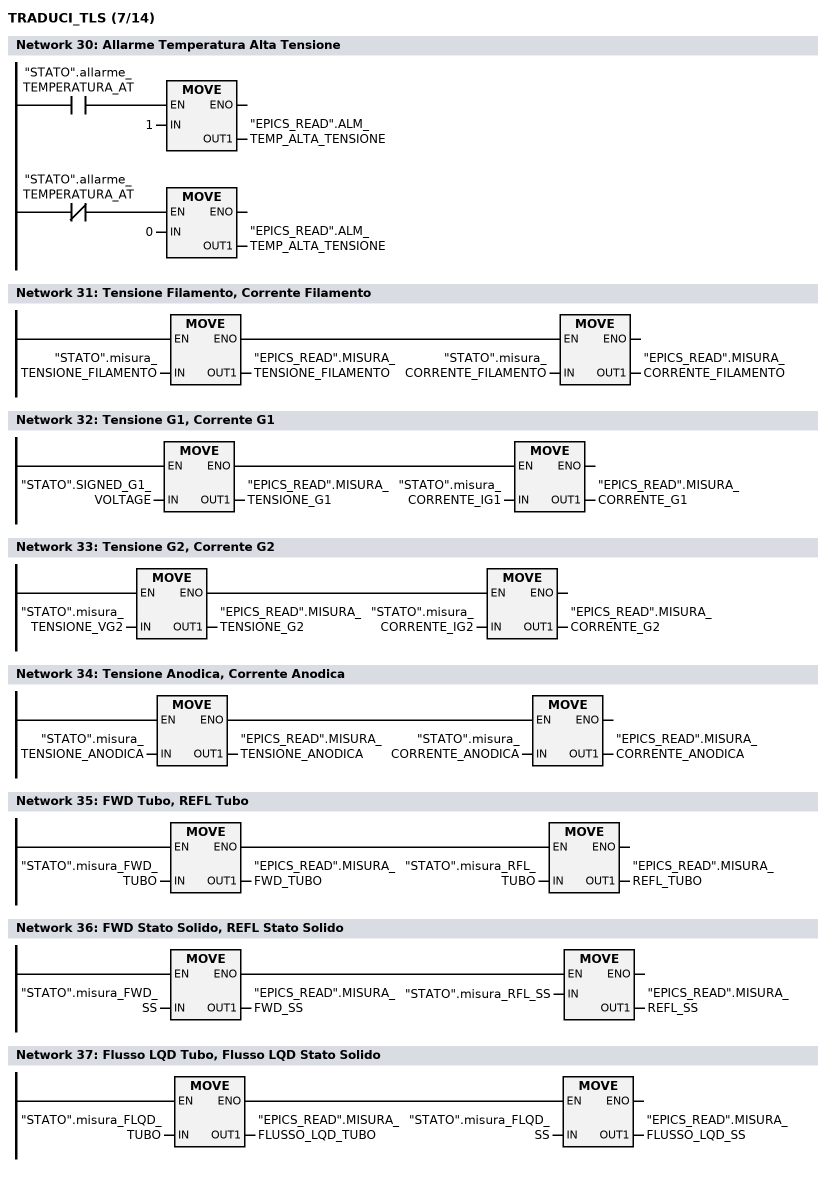
   RUNG wire#powerrail
      Contact( "STATO".allarme_TEMPERATURA_AT )
      Move(in := 1, out1 => "EPICS_READ".ALM_TEMP_ALTA_TENSIONE)
   END_RUNG
   RUNG wire#powerrail
      I_Contact( "STATO".allarme_TEMPERATURA_AT )
      Move(in := 0, out1 => "EPICS_READ".ALM_TEMP_ALTA_TENSIONE)
   END_RUNG
   // the same network as SCL:
   IF "STATO".allarme_TEMPERATURA_AT THEN "EPICS_READ".ALM_TEMP_ALTA_TENSIONE := 1; END_IF;
   IF NOT "STATO".allarme_TEMPERATURA_AT THEN "EPICS_READ".ALM_TEMP_ALTA_TENSIONE := 0; END_IF;
END_REGION

REGION Network 31: Tensione Filamento, Corrente Filamento
   RUNG wire#powerrail
      Move(in := "STATO".misura_TENSIONE_FILAMENTO, out1 => "EPICS_READ".MISURA_TENSIONE_FILAMENTO)
      Move(in := "STATO".misura_CORRENTE_FILAMENTO, out1 => "EPICS_READ".MISURA_CORRENTE_FILAMENTO)
   END_RUNG
   // the same network as SCL:
   "EPICS_READ".MISURA_TENSIONE_FILAMENTO := "STATO".misura_TENSIONE_FILAMENTO;
   "EPICS_READ".MISURA_CORRENTE_FILAMENTO := "STATO".misura_CORRENTE_FILAMENTO;
END_REGION

REGION Network 32: Tensione G1, Corrente G1
   RUNG wire#powerrail
      Move(in := "STATO".SIGNED_G1_VOLTAGE, out1 => "EPICS_READ".MISURA_TENSIONE_G1)
      Move(in := "STATO".misura_CORRENTE_IG1, out1 => "EPICS_READ".MISURA_CORRENTE_G1)
   END_RUNG
   // the same network as SCL:
   "EPICS_READ".MISURA_TENSIONE_G1 := "STATO".SIGNED_G1_VOLTAGE;
   "EPICS_READ".MISURA_CORRENTE_G1 := "STATO".misura_CORRENTE_IG1;
END_REGION

REGION Network 33: Tensione G2, Corrente G2
   RUNG wire#powerrail
      Move(in := "STATO".misura_TENSIONE_VG2, out1 => "EPICS_READ".MISURA_TENSIONE_G2)
      Move(in := "STATO".misura_CORRENTE_IG2, out1 => "EPICS_READ".MISURA_CORRENTE_G2)
   END_RUNG
   // the same network as SCL:
   "EPICS_READ".MISURA_TENSIONE_G2 := "STATO".misura_TENSIONE_VG2;
   "EPICS_READ".MISURA_CORRENTE_G2 := "STATO".misura_CORRENTE_IG2;
END_REGION

REGION Network 34: Tensione Anodica, Corrente Anodica
   RUNG wire#powerrail
      Move(in := "STATO".misura_TENSIONE_ANODICA, out1 => "EPICS_READ".MISURA_TENSIONE_ANODICA)
      Move(in := "STATO".misura_CORRENTE_ANODICA, out1 => "EPICS_READ".MISURA_CORRENTE_ANODICA)
   END_RUNG
   // the same network as SCL:
   "EPICS_READ".MISURA_TENSIONE_ANODICA := "STATO".misura_TENSIONE_ANODICA;
   "EPICS_READ".MISURA_CORRENTE_ANODICA := "STATO".misura_CORRENTE_ANODICA;
END_REGION

REGION Network 35: FWD Tubo, REFL Tubo
   RUNG wire#powerrail
      Move(in := "STATO".misura_FWD_TUBO, out1 => "EPICS_READ".MISURA_FWD_TUBO)
      Move(in := "STATO".misura_RFL_TUBO, out1 => "EPICS_READ".MISURA_REFL_TUBO)
   END_RUNG
   // the same network as SCL:
   "EPICS_READ".MISURA_FWD_TUBO := "STATO".misura_FWD_TUBO;
   "EPICS_READ".MISURA_REFL_TUBO := "STATO".misura_RFL_TUBO;
END_REGION

REGION Network 36: FWD Stato Solido, REFL Stato Solido
   RUNG wire#powerrail
      Move(in := "STATO".misura_FWD_SS, out1 => "EPICS_READ".MISURA_FWD_SS)
      Move(in := "STATO".misura_RFL_SS, out1 => "EPICS_READ".MISURA_REFL_SS)
   END_RUNG
   // the same network as SCL:
   "EPICS_READ".MISURA_FWD_SS := "STATO".misura_FWD_SS;
   "EPICS_READ".MISURA_REFL_SS := "STATO".misura_RFL_SS;
END_REGION

REGION Network 37: Flusso LQD Tubo, Flusso LQD Stato Solido
   RUNG wire#powerrail
      Move(in := "STATO".misura_FLQD_TUBO, out1 => "EPICS_READ".MISURA_FLUSSO_LQD_TUBO)
      Move(in := "STATO".misura_FLQD_SS, out1 => "EPICS_READ".MISURA_FLUSSO_LQD_SS)
   END_RUNG
   // the same network as SCL:
   "EPICS_READ".MISURA_FLUSSO_LQD_TUBO := "STATO".misura_FLQD_TUBO;
   "EPICS_READ".MISURA_FLUSSO_LQD_SS := "STATO".misura_FLQD_SS;
END_REGION

REGION Network 38: Temperature LQD IN/OUT Tubo, Stato Solido